REGION Network 10: Stacker General Alarm
   RUNG wire#powerrail
      { S7_Templates := "SrcType := Word" } EQ_Contact(in1 := "DB3_FAULTS".Alarm_Safety_S, in2 := 0)
      { S7_Templates := "SrcType := Word" } EQ_Contact(in1 := "DB3_FAULTS".Alarm_Safety_SN, in2 := 0)
      { S7_Templates := "SrcType := Word" } EQ_Contact(in1 := "DB3_FAULTS".Alarm_Safety_Z2, in2 := 0)
      { S7_Templates := "SrcType := Word" } EQ_Contact(in1 := "DB3_FAULTS".Alarm_Stacker, in2 := 0)
      { S7_Templates := "SrcType := Word" } EQ_Contact(in1 := "DB3_FAULTS".Alarm_General_S, in2 := 0)
      { S7_Templates := "SrcType := Word" } EQ_Contact(in1 := "DB3_FAULTS".Alarm_CD2, in2 := 0)
      { S7_Templates := "SrcType := Word" } EQ_Contact(in1 := "DB3_FAULTS".Alarm_CD1, in2 := 0)
      Coil( #NoAlmAny )
   END_RUNG
   RUNG wire#powerrail
      Contact( #NoAlmAny )
      { S7_Templates := "SrcType := Word" } EQ_Contact(in1 := "s".f[1].almw, in2 := 0)
      { S7_Templates := "SrcType := Word" } EQ_Contact(in1 := "s".f[2].almw, in2 := 0)
      { S7_Templates := "SrcType := Word" } EQ_Contact(in1 := "s".f[3].almw, in2 := 0)
      { S7_Templates := "SrcType := Word" } EQ_Contact(in1 := "s".f[4].almw, in2 := 0)
      { S7_Templates := "SrcType := Word" } EQ_Contact(in1 := "s".f[5].almw, in2 := 0)
      Coil( #NoAlmAny )
   END_RUNG
   RUNG wire#powerrail
      Contact( #NoAlmAny )
      { S7_Templates := "SrcType := Word" } EQ_Contact(in1 := "O".S_Alm_Stack_Dwn, in2 := 0)
      { S7_Templates := "SrcType := Word" } EQ_Contact(in1 := "O".S_Alm_Stack_Mid, in2 := 0)
      { S7_Templates := "SrcType := Word" } EQ_Contact(in1 := "O".S_Alm_Stack_Up, in2 := 0)
      { S7_Templates := "SrcType := Word" } EQ_Contact(in1 := "O".Centror_A.AlarmW, in2 := 0)
      { S7_Templates := "SrcType := Word" } EQ_Contact(in1 := "O".FurcaStacker.AlarmW, in2 := 0)
      I_Contact( "DB2_WORK_BITS".Stacker_Handler.Output.oAlarmForks )
      I_Contact( "DB2_WORK_BITS".Stacker_Handler.Output.oAlarmPosition )
      Coil( #NoAlmAny )
   END_RUNG
   RUNG wire#powerrail
      I_Contact( #NoAlmAny )
      I_Contact( "x"."b"[16] )
      Coil( "Gen".S_AlarmAny )
   END_RUNG
   // the same network as SCL:
   #NoAlmAny := ("DB3_FAULTS".Alarm_Safety_S = 0) AND ("DB3_FAULTS".Alarm_Safety_SN = 0) AND ("DB3_FAULTS".Alarm_Safety_Z2 = 0) AND ("DB3_FAULTS".Alarm_Stacker = 0) AND ("DB3_FAULTS".Alarm_General_S = 0) AND ("DB3_FAULTS".Alarm_CD2 = 0) AND ("DB3_FAULTS".Alarm_CD1 = 0);
   #NoAlmAny := #NoAlmAny AND ("s".f[1].almw = 0) AND ("s".f[2].almw = 0) AND ("s".f[3].almw = 0) AND ("s".f[4].almw = 0) AND ("s".f[5].almw = 0);
   #NoAlmAny := #NoAlmAny AND ("O".S_Alm_Stack_Dwn = 0) AND ("O".S_Alm_Stack_Mid = 0) AND ("O".S_Alm_Stack_Up = 0) AND ("O".Centror_A.AlarmW = 0) AND ("O".FurcaStacker.AlarmW = 0) AND NOT "DB2_WORK_BITS".Stacker_Handler.Output.oAlarmForks AND NOT "DB2_WORK_BITS".Stacker_Handler.Output.oAlarmPosition;
   "Gen".S_AlarmAny := NOT #NoAlmAny AND NOT "x"."b"[16];
END_REGION

REGION Network 11: Stacker_New General Alarm
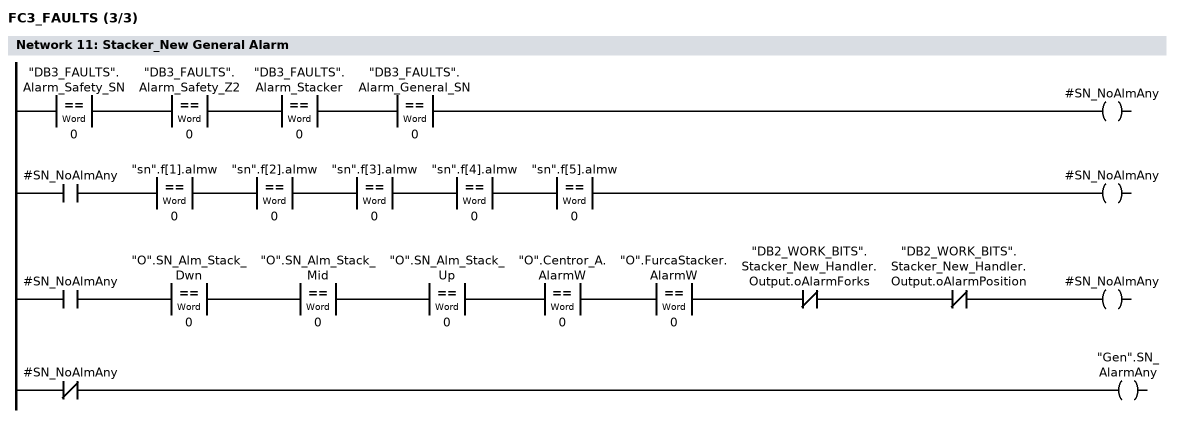
   RUNG wire#powerrail
      { S7_Templates := "SrcType := Word" } EQ_Contact(in1 := "DB3_FAULTS".Alarm_Safety_SN, in2 := 0)
      { S7_Templates := "SrcType := Word" } EQ_Contact(in1 := "DB3_FAULTS".Alarm_Safety_Z2, in2 := 0)
      { S7_Templates := "SrcType := Word" } EQ_Contact(in1 := "DB3_FAULTS".Alarm_Stacker, in2 := 0)
      { S7_Templates := "SrcType := Word" } EQ_Contact(in1 := "DB3_FAULTS".Alarm_General_SN, in2 := 0)
      Coil( #SN_NoAlmAny )
   END_RUNG
   RUNG wire#powerrail
      Contact( #SN_NoAlmAny )
      { S7_Templates := "SrcType := Word" } EQ_Contact(in1 := "sn".f[1].almw, in2 := 0)
      { S7_Templates := "SrcType := Word" } EQ_Contact(in1 := "sn".f[2].almw, in2 := 0)
      { S7_Templates := "SrcType := Word" } EQ_Contact(in1 := "sn".f[3].almw, in2 := 0)
      { S7_Templates := "SrcType := Word" } EQ_Contact(in1 := "sn".f[4].almw, in2 := 0)
      { S7_Templates := "SrcType := Word" } EQ_Contact(in1 := "sn".f[5].almw, in2 := 0)
      Coil( #SN_NoAlmAny )
   END_RUNG
   RUNG wire#powerrail
      Contact( #SN_NoAlmAny )
      { S7_Templates := "SrcType := Word" } EQ_Contact(in1 := "O".SN_Alm_Stack_Dwn, in2 := 0)
      { S7_Templates := "SrcType := Word" } EQ_Contact(in1 := "O".SN_Alm_Stack_Mid, in2 := 0)
      { S7_Templates := "SrcType := Word" } EQ_Contact(in1 := "O".SN_Alm_Stack_Up, in2 := 0)
      { S7_Templates := "SrcType := Word" } EQ_Contact(in1 := "O".Centror_A.AlarmW, in2 := 0)
      { S7_Templates := "SrcType := Word" } EQ_Contact(in1 := "O".FurcaStacker.AlarmW, in2 := 0)
      I_Contact( "DB2_WORK_BITS".Stacker_New_Handler.Output.oAlarmForks )
      I_Contact( "DB2_WORK_BITS".Stacker_New_Handler.Output.oAlarmPosition )
      Coil( #SN_NoAlmAny )
   END_RUNG
   RUNG wire#powerrail
      I_Contact( #SN_NoAlmAny )
      Coil( "Gen".SN_AlarmAny )
   END_RUNG
   // the same network as SCL:
   #SN_NoAlmAny := ("DB3_FAULTS".Alarm_Safety_SN = 0) AND ("DB3_FAULTS".Alarm_Safety_Z2 = 0) AND ("DB3_FAULTS".Alarm_Stacker = 0) AND ("DB3_FAULTS".Alarm_General_SN = 0);
   #SN_NoAlmAny := #SN_NoAlmAny AND ("sn".f[1].almw = 0) AND ("sn".f[2].almw = 0) AND ("sn".f[3].almw = 0) AND ("sn".f[4].almw = 0) AND ("sn".f[5].almw = 0);
   #SN_NoAlmAny := #SN_NoAlmAny AND ("O".SN_Alm_Stack_Dwn = 0) AND ("O".SN_Alm_Stack_Mid = 0) AND ("O".SN_Alm_Stack_Up = 0) AND ("O".Centror_A.AlarmW = 0) AND ("O".FurcaStacker.AlarmW = 0) AND NOT "DB2_WORK_BITS".Stacker_New_Handler.Output.oAlarmForks AND NOT "DB2_WORK_BITS".Stacker_New_Handler.Output.oAlarmPosition;
   "Gen".SN_AlarmAny := NOT #SN_NoAlmAny;
END_REGION
END_FUNCTION

FUNCTION "FC6_OUTPUTS" : Void   // FC6, LAD
{ S7_Optimized_Access := 'TRUE' }
VERSION : 0.1
   VAR_TEMP
      S_bsy : Bool;
      S_bsg : Bool;
      S_bsr : Bool;
      S_bsgc : Bool;
      cfo1 : Bool;
      cfo2 : Bool;
      cfo3 : Bool;
      cfA : Bool;
      SN_bsr : Bool;
      SN_bsy : Bool;
      SN_bsgc : Bool;
      SN_bsg : Bool;
      SN_cfo1 : Bool;
      SN_cfo2 : Bool;
      SN_cfo3 : Bool;
      SN_cfA : Bool;
   END_VAR
   VAR_TEMP   // added for the SCL form of the ladder/FBD networks
      _w1 : Bool;
   END_VAR
BEGIN

REGION Network 1: Stacking_New VFD Input Conveyor
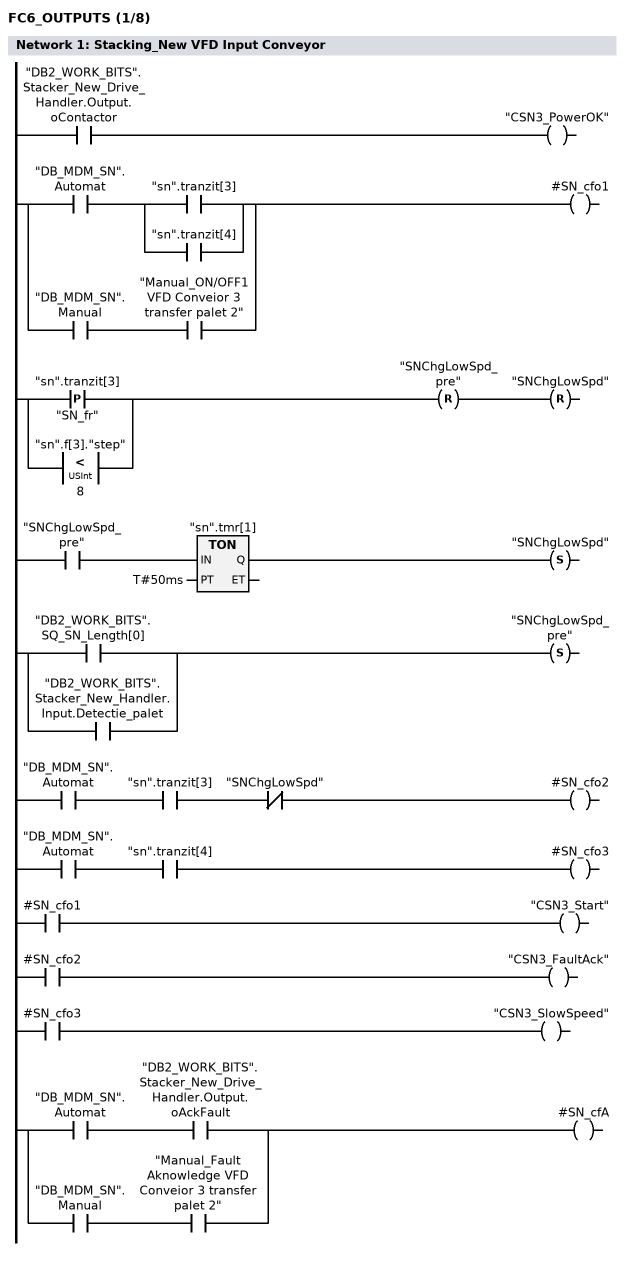
   "CSN3_PowerOK" := "DB2_WORK_BITS".Stacker_New_Drive_Handler.Output.oContactor;
   #SN_cfo1 := ("DB_MDM_SN".Automat AND ("sn".tranzit[3] OR "sn".tranzit[4])) OR ("DB_MDM_SN".Manual AND "Manual_ON/OFF1 VFD Conveior 3 transfer palet 2");
   #_w1 := "sn".tranzit[3] AND NOT "SN_fr";   // rising edge of "sn".tranzit[3]
   "SN_fr" := "sn".tranzit[3];
   IF #_w1 OR ("sn".f[3]."step" < 8) THEN
       "SNChgLowSpd_pre" := FALSE;
       "SNChgLowSpd" := FALSE;
   END_IF;
   "sn".tmr[1].TON(IN := "SNChgLowSpd_pre", PT := T#50ms);
   IF "sn".tmr[1].Q THEN "SNChgLowSpd" := TRUE; END_IF;
   IF "DB2_WORK_BITS".SQ_SN_Length[0] OR "DB2_WORK_BITS".Stacker_New_Handler.Input.Detectie_palet THEN
       "SNChgLowSpd_pre" := TRUE;
   END_IF;
   #SN_cfo2 := "DB_MDM_SN".Automat AND "sn".tranzit[3] AND NOT "SNChgLowSpd";
   #SN_cfo3 := "DB_MDM_SN".Automat AND "sn".tranzit[4];
   "CSN3_Start" := #SN_cfo1;
   "CSN3_FaultAck" := #SN_cfo2;
   "CSN3_SlowSpeed" := #SN_cfo3;
   #SN_cfA := ("DB_MDM_SN".Automat AND "DB2_WORK_BITS".Stacker_New_Drive_Handler.Output.oAckFault) OR ("DB_MDM_SN".Manual AND "Manual_Fault Aknowledge VFD Conveior 3 transfer palet 2");
END_REGION

REGION Network 2: Stacking_New VFD Output Conveyor
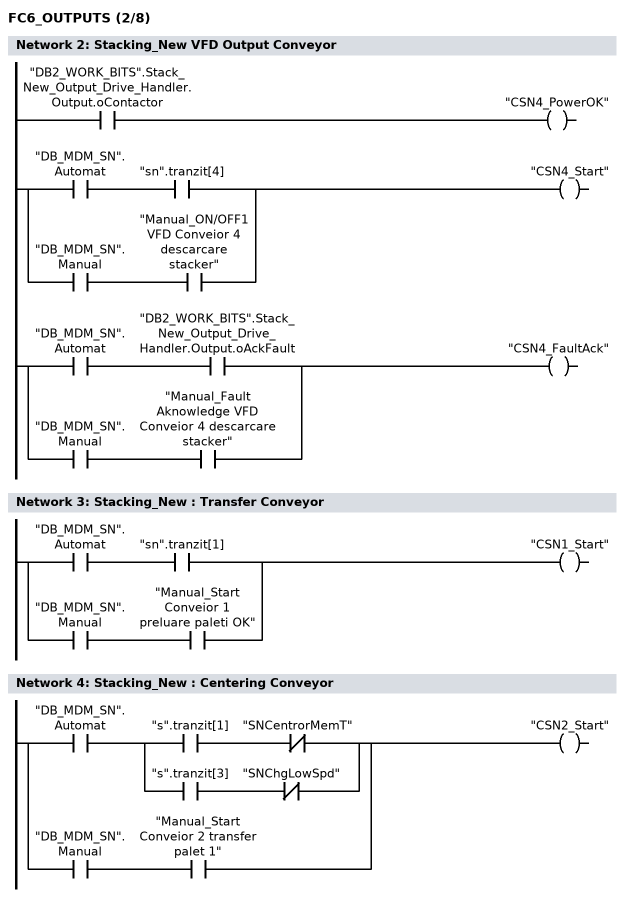
   RUNG wire#powerrail
      Contact( "DB2_WORK_BITS".Stack_New_Output_Drive_Handler.Output.oContactor )
      Coil( "CSN4_PowerOK" )
   END_RUNG
   RUNG wire#powerrail
      Contact( "DB_MDM_SN".Automat )
      Contact( "sn".tranzit[4] )
      wire#w1
      Coil( "CSN4_Start" )
   END_RUNG
   RUNG wire#powerrail
      Contact( "DB_MDM_SN".Manual )
      Contact( "Manual_ON/OFF1 VFD Conveior 4 descarcare stacker" )
   END_RUNG wire#w1
   RUNG wire#powerrail
      Contact( "DB_MDM_SN".Automat )
      Contact( "DB2_WORK_BITS".Stack_New_Output_Drive_Handler.Output.oAckFault )
      wire#w2
      Coil( "CSN4_FaultAck" )
   END_RUNG
   RUNG wire#powerrail
      Contact( "DB_MDM_SN".Manual )
      Contact( "Manual_Fault Aknowledge VFD Conveior 4 descarcare stacker" )
   END_RUNG wire#w2
   // the same network as SCL:
   "CSN4_PowerOK" := "DB2_WORK_BITS".Stack_New_Output_Drive_Handler.Output.oContactor;
   "CSN4_Start" := ("DB_MDM_SN".Automat AND "sn".tranzit[4]) OR ("DB_MDM_SN".Manual AND "Manual_ON/OFF1 VFD Conveior 4 descarcare stacker");
   "CSN4_FaultAck" := ("DB_MDM_SN".Automat AND "DB2_WORK_BITS".Stack_New_Output_Drive_Handler.Output.oAckFault) OR ("DB_MDM_SN".Manual AND "Manual_Fault Aknowledge VFD Conveior 4 descarcare stacker");
END_REGION

REGION Network 3: Stacking_New : Transfer Conveyor
   RUNG wire#powerrail
      Contact( "DB_MDM_SN".Automat )
      Contact( "sn".tranzit[1] )
      wire#w1
      Coil( "CSN1_Start" )
   END_RUNG
   RUNG wire#powerrail
      Contact( "DB_MDM_SN".Manual )
      Contact( "Manual_Start Conveior 1 preluare paleti OK" )
   END_RUNG wire#w1
   // the same network as SCL:
   "CSN1_Start" := ("DB_MDM_SN".Automat AND "sn".tranzit[1]) OR ("DB_MDM_SN".Manual AND "Manual_Start Conveior 1 preluare paleti OK");
END_REGION

REGION Network 4: Stacking_New : Centering Conveyor
   RUNG wire#powerrail
      Contact( "DB_MDM_SN".Automat )
      wire#w1
      Contact( "s".tranzit[1] )
      I_Contact( "SNCentrorMemT" )
      wire#w2
      Coil( "CSN2_Start" )
   END_RUNG
   RUNG wire#w1
      Contact( "s".tranzit[3] )
      I_Contact( "SNChgLowSpd" )
   END_RUNG wire#w2
   RUNG wire#powerrail
      Contact( "DB_MDM_SN".Manual )
      Contact( "Manual_Start Conveior 2 transfer palet 1" )
   END_RUNG wire#w2
   // the same network as SCL:
   "CSN2_Start" := ("DB_MDM_SN".Automat AND (("s".tranzit[1] AND NOT "SNCentrorMemT") OR ("s".tranzit[3] AND NOT "SNChgLowSpd"))) OR ("DB_MDM_SN".Manual AND "Manual_Start Conveior 2 transfer palet 1");
END_REGION

REGION Network 5: Stacking : VFD Input Conveyor
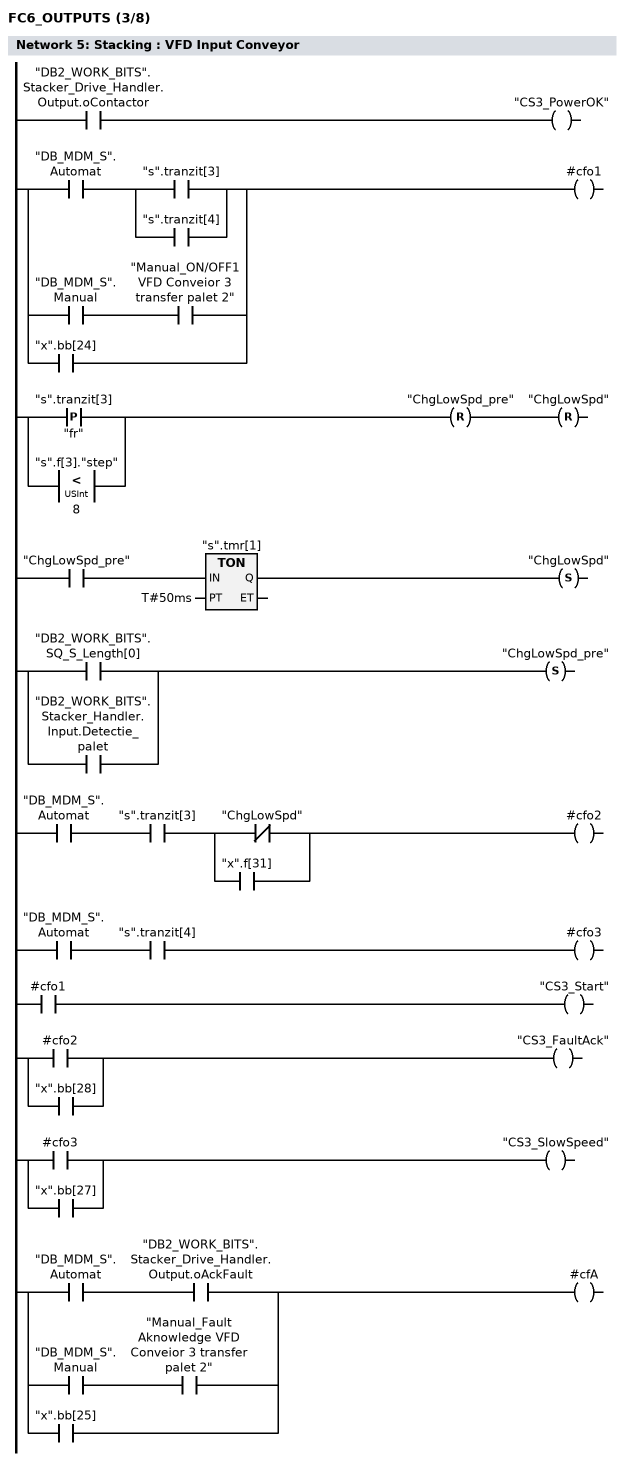
   "CS3_PowerOK" := "DB2_WORK_BITS".Stacker_Drive_Handler.Output.oContactor;
   #cfo1 := ("DB_MDM_S".Automat AND ("s".tranzit[3] OR "s".tranzit[4])) OR ("DB_MDM_S".Manual AND "Manual_ON/OFF1 VFD Conveior 3 transfer palet 2") OR "x".bb[24];
   #_w1 := "s".tranzit[3] AND NOT "fr";   // rising edge of "s".tranzit[3]
   "fr" := "s".tranzit[3];
   IF #_w1 OR ("s".f[3]."step" < 8) THEN
       "ChgLowSpd_pre" := FALSE;
       "ChgLowSpd" := FALSE;
   END_IF;
   "s".tmr[1].TON(IN := "ChgLowSpd_pre", PT := T#50ms);
   IF "s".tmr[1].Q THEN "ChgLowSpd" := TRUE; END_IF;
   IF "DB2_WORK_BITS".SQ_S_Length[0] OR "DB2_WORK_BITS".Stacker_Handler.Input.Detectie_palet THEN
       "ChgLowSpd_pre" := TRUE;
   END_IF;
   #cfo2 := "DB_MDM_S".Automat AND "s".tranzit[3] AND (NOT "ChgLowSpd" OR "x".f[31]);
   #cfo3 := "DB_MDM_S".Automat AND "s".tranzit[4];
   "CS3_Start" := #cfo1;
   "CS3_FaultAck" := #cfo2 OR "x".bb[28];
   "CS3_SlowSpeed" := #cfo3 OR "x".bb[27];
   #cfA := ("DB_MDM_S".Automat AND "DB2_WORK_BITS".Stacker_Drive_Handler.Output.oAckFault) OR ("DB_MDM_S".Manual AND "Manual_Fault Aknowledge VFD Conveior 3 transfer palet 2") OR "x".bb[25];
END_REGION

REGION Network 6: Stacking : VFD Output Conveyor
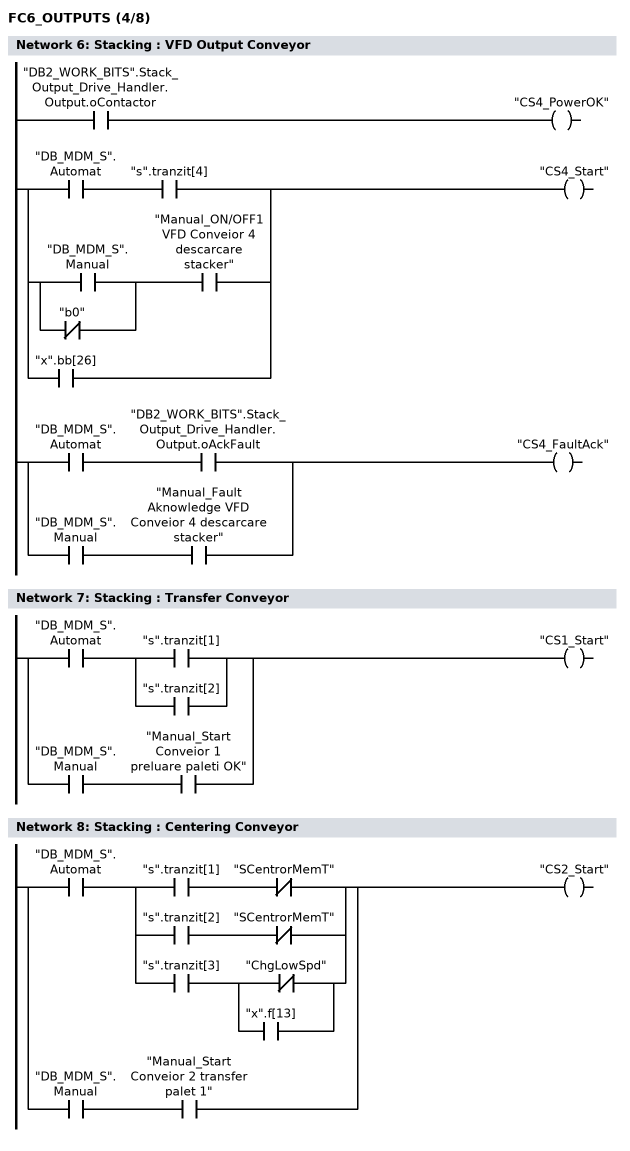
   RUNG wire#powerrail
      Contact( "DB2_WORK_BITS".Stack_Output_Drive_Handler.Output.oContactor )
      Coil( "CS4_PowerOK" )
   END_RUNG
   RUNG wire#powerrail
      Contact( "DB_MDM_S".Automat )
      Contact( "s".tranzit[4] )
      wire#w1
      Coil( "CS4_Start" )
   END_RUNG
   RUNG wire#powerrail
      Contact( "DB_MDM_S".Manual )
      wire#w2
      Contact( "Manual_ON/OFF1 VFD Conveior 4 descarcare stacker" )
   END_RUNG wire#w1
   RUNG wire#powerrail
      I_Contact( "b0" )
   END_RUNG wire#w2
   RUNG wire#powerrail
      Contact( "x".bb[26] )
   END_RUNG wire#w1
   RUNG wire#powerrail
      Contact( "DB_MDM_S".Automat )
      Contact( "DB2_WORK_BITS".Stack_Output_Drive_Handler.Output.oAckFault )
      wire#w3
      Coil( "CS4_FaultAck" )
   END_RUNG
   RUNG wire#powerrail
      Contact( "DB_MDM_S".Manual )
      Contact( "Manual_Fault Aknowledge VFD Conveior 4 descarcare stacker" )
   END_RUNG wire#w3
   // the same network as SCL:
   "CS4_PowerOK" := "DB2_WORK_BITS".Stack_Output_Drive_Handler.Output.oContactor;
   "CS4_Start" := ("DB_MDM_S".Automat AND "s".tranzit[4]) OR (("DB_MDM_S".Manual OR NOT "b0") AND "Manual_ON/OFF1 VFD Conveior 4 descarcare stacker") OR "x".bb[26];
   "CS4_FaultAck" := ("DB_MDM_S".Automat AND "DB2_WORK_BITS".Stack_Output_Drive_Handler.Output.oAckFault) OR ("DB_MDM_S".Manual AND "Manual_Fault Aknowledge VFD Conveior 4 descarcare stacker");
END_REGION

REGION Network 7: Stacking : Transfer Conveyor
   RUNG wire#powerrail
      Contact( "DB_MDM_S".Automat )
      wire#w1
      Contact( "s".tranzit[1] )
      wire#w2
      Coil( "CS1_Start" )
   END_RUNG
   RUNG wire#w1
      Contact( "s".tranzit[2] )
   END_RUNG wire#w2
   RUNG wire#powerrail
      Contact( "DB_MDM_S".Manual )
      Contact( "Manual_Start Conveior 1 preluare paleti OK" )
   END_RUNG wire#w2
   // the same network as SCL:
   "CS1_Start" := ("DB_MDM_S".Automat AND ("s".tranzit[1] OR "s".tranzit[2])) OR ("DB_MDM_S".Manual AND "Manual_Start Conveior 1 preluare paleti OK");
END_REGION

REGION Network 8: Stacking : Centering Conveyor
   RUNG wire#powerrail
      Contact( "DB_MDM_S".Automat )
      wire#w1
      Contact( "s".tranzit[1] )
      I_Contact( "SCentrorMemT" )
      wire#w2
      Coil( "CS2_Start" )
   END_RUNG
   RUNG wire#w1
      Contact( "s".tranzit[2] )
      I_Contact( "SCentrorMemT" )
   END_RUNG wire#w2
   RUNG wire#w1
      Contact( "s".tranzit[3] )
      wire#w3
      I_Contact( "ChgLowSpd" )
   END_RUNG wire#w2
   RUNG wire#w3
      Contact( "x".f[13] )
   END_RUNG wire#w2
   RUNG wire#powerrail
      Contact( "DB_MDM_S".Manual )
      Contact( "Manual_Start Conveior 2 transfer palet 1" )
   END_RUNG wire#w2
   // the same network as SCL:
   "CS2_Start" := ("DB_MDM_S".Automat AND (("s".tranzit[1] AND NOT "SCentrorMemT") OR ("s".tranzit[2] AND NOT "SCentrorMemT") OR ("s".tranzit[3] AND (NOT "ChgLowSpd" OR "x".f[13])))) OR ("DB_MDM_S".Manual AND "Manual_Start Conveior 2 transfer palet 1");
END_REGION

REGION Network 9: Stacking_New : Comanda SoftStart Power ON
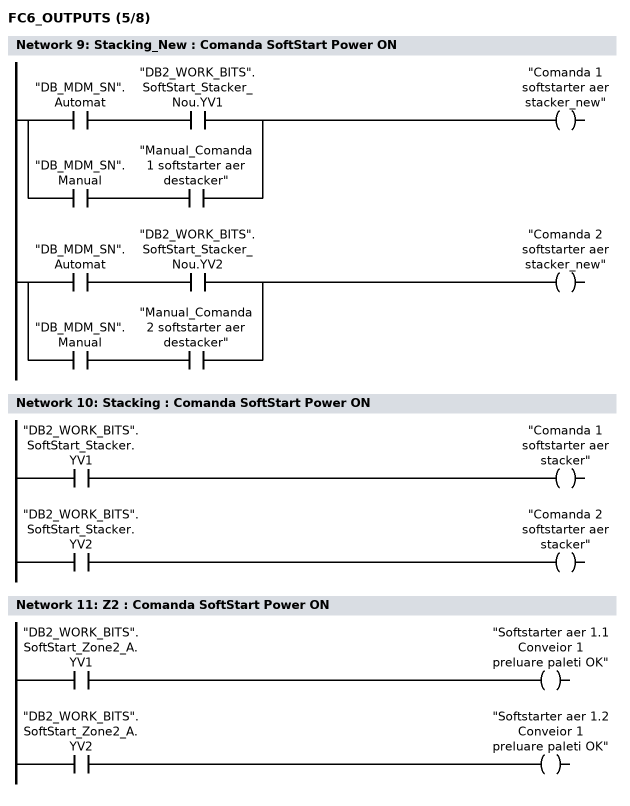
   RUNG wire#powerrail
      Contact( "DB_MDM_SN".Automat )
      Contact( "DB2_WORK_BITS".SoftStart_Stacker_Nou.YV1 )
      wire#w1
      Coil( "Comanda 1 softstarter aer stacker_new" )
   END_RUNG
   RUNG wire#powerrail
      Contact( "DB_MDM_SN".Manual )
      Contact( "Manual_Comanda 1 softstarter aer destacker" )
   END_RUNG wire#w1
   RUNG wire#powerrail
      Contact( "DB_MDM_SN".Automat )
      Contact( "DB2_WORK_BITS".SoftStart_Stacker_Nou.YV2 )
      wire#w2
      Coil( "Comanda 2 softstarter aer stacker_new" )
   END_RUNG
   RUNG wire#powerrail
      Contact( "DB_MDM_SN".Manual )
      Contact( "Manual_Comanda 2 softstarter aer destacker" )
   END_RUNG wire#w2
   // the same network as SCL:
   "Comanda 1 softstarter aer stacker_new" := ("DB_MDM_SN".Automat AND "DB2_WORK_BITS".SoftStart_Stacker_Nou.YV1) OR ("DB_MDM_SN".Manual AND "Manual_Comanda 1 softstarter aer destacker");
   "Comanda 2 softstarter aer stacker_new" := ("DB_MDM_SN".Automat AND "DB2_WORK_BITS".SoftStart_Stacker_Nou.YV2) OR ("DB_MDM_SN".Manual AND "Manual_Comanda 2 softstarter aer destacker");
END_REGION

REGION Network 10: Stacking : Comanda SoftStart Power ON
   RUNG wire#powerrail
      Contact( "DB2_WORK_BITS".SoftStart_Stacker.YV1 )
      Coil( "Comanda 1 softstarter aer stacker" )
   END_RUNG
   RUNG wire#powerrail
      Contact( "DB2_WORK_BITS".SoftStart_Stacker.YV2 )
      Coil( "Comanda 2 softstarter aer stacker" )
   END_RUNG
   // the same network as SCL:
   "Comanda 1 softstarter aer stacker" := "DB2_WORK_BITS".SoftStart_Stacker.YV1;
   "Comanda 2 softstarter aer stacker" := "DB2_WORK_BITS".SoftStart_Stacker.YV2;
END_REGION

REGION Network 11: Z2 : Comanda SoftStart Power ON
   RUNG wire#powerrail
      Contact( "DB2_WORK_BITS".SoftStart_Zone2_A.YV1 )
      Coil( "Softstarter aer 1.1 Conveior 1 preluare paleti OK" )
   END_RUNG
   RUNG wire#powerrail
      Contact( "DB2_WORK_BITS".SoftStart_Zone2_A.YV2 )
      Coil( "Softstarter aer 1.2 Conveior 1 preluare paleti OK" )
   END_RUNG
   // the same network as SCL:
   "Softstarter aer 1.1 Conveior 1 preluare paleti OK" := "DB2_WORK_BITS".SoftStart_Zone2_A.YV1;
   "Softstarter aer 1.2 Conveior 1 preluare paleti OK" := "DB2_WORK_BITS".SoftStart_Zone2_A.YV2;
END_REGION

REGION Network 12: Rearm safety
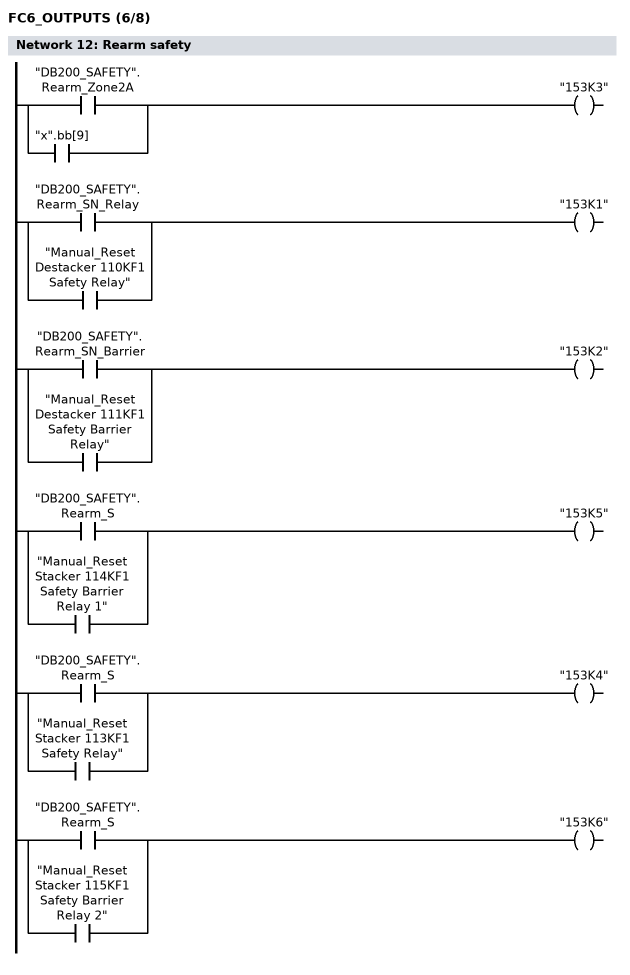
   RUNG wire#powerrail
      Contact( "DB200_SAFETY".Rearm_Zone2A )
      wire#w1
      Coil( "153K3" )
   END_RUNG
   RUNG wire#powerrail
      Contact( "x".bb[9] )
   END_RUNG wire#w1
   RUNG wire#powerrail
      Contact( "DB200_SAFETY".Rearm_SN_Relay )
      wire#w2
      Coil( "153K1" )
   END_RUNG
   RUNG wire#powerrail
      Contact( "Manual_Reset Destacker 110KF1 Safety Relay" )
   END_RUNG wire#w2
   RUNG wire#powerrail
      Contact( "DB200_SAFETY".Rearm_SN_Barrier )
      wire#w3
      Coil( "153K2" )
   END_RUNG
   RUNG wire#powerrail
      Contact( "Manual_Reset Destacker 111KF1 Safety Barrier Relay" )
   END_RUNG wire#w3
   RUNG wire#powerrail
      Contact( "DB200_SAFETY".Rearm_S )
      wire#w4
      Coil( "153K5" )
   END_RUNG
   RUNG wire#powerrail
      Contact( "Manual_Reset Stacker 114KF1 Safety Barrier Relay 1" )
   END_RUNG wire#w4
   RUNG wire#powerrail
      Contact( "DB200_SAFETY".Rearm_S )
      wire#w5
      Coil( "153K4" )
   END_RUNG
   RUNG wire#powerrail
      Contact( "Manual_Reset Stacker 113KF1 Safety Relay" )
   END_RUNG wire#w5
   RUNG wire#powerrail
      Contact( "DB200_SAFETY".Rearm_S )
      wire#w6
      Coil( "153K6" )
   END_RUNG
   RUNG wire#powerrail
      Contact( "Manual_Reset Stacker 115KF1 Safety Barrier Relay 2" )
   END_RUNG wire#w6
   // the same network as SCL:
   "153K3" := "DB200_SAFETY".Rearm_Zone2A OR "x".bb[9];
   "153K1" := "DB200_SAFETY".Rearm_SN_Relay OR "Manual_Reset Destacker 110KF1 Safety Relay";
   "153K2" := "DB200_SAFETY".Rearm_SN_Barrier OR "Manual_Reset Destacker 111KF1 Safety Barrier Relay";
   "153K5" := "DB200_SAFETY".Rearm_S OR "Manual_Reset Stacker 114KF1 Safety Barrier Relay 1";
   "153K4" := "DB200_SAFETY".Rearm_S OR "Manual_Reset Stacker 113KF1 Safety Relay";
   "153K6" := "DB200_SAFETY".Rearm_S OR "Manual_Reset Stacker 115KF1 Safety Barrier Relay 2";
END_REGION

REGION Network 13: Stacking : Control Balize
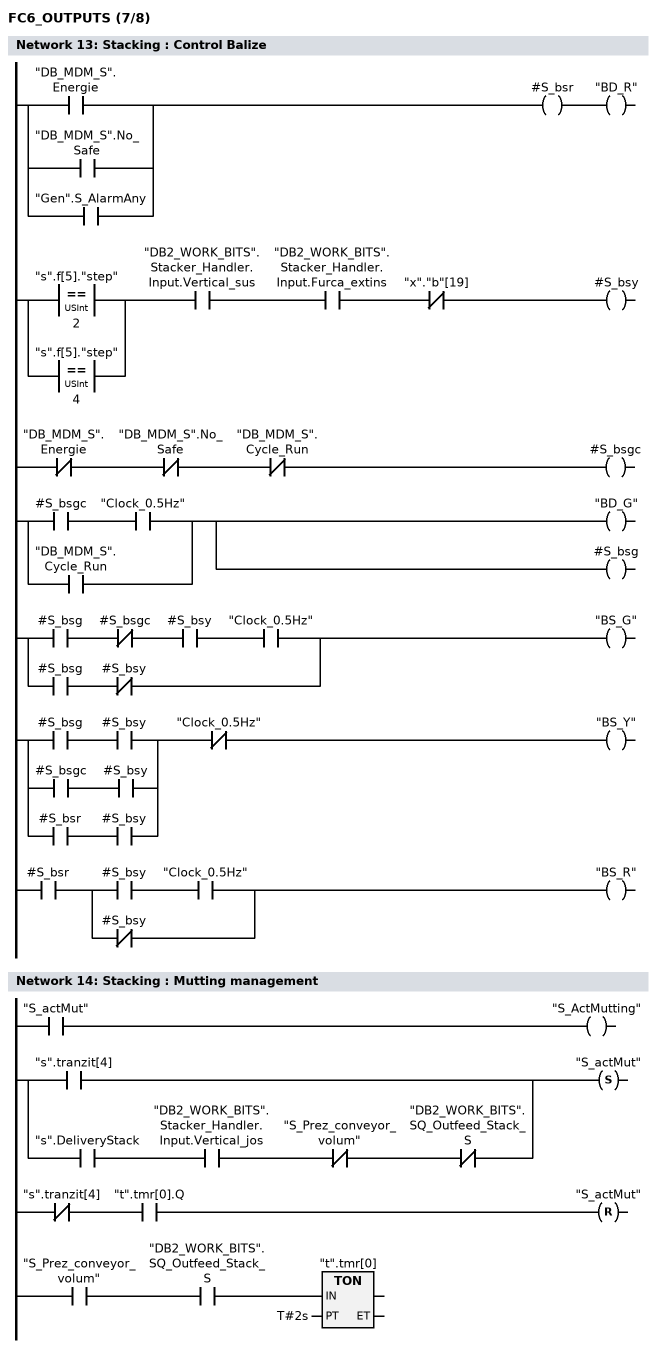
   RUNG wire#powerrail
      Contact( "DB_MDM_S".Energie )
      wire#w1
      Coil( #S_bsr )
      Coil( "BD_R" )
   END_RUNG
   RUNG wire#powerrail
      Contact( "DB_MDM_S".No_Safe )
   END_RUNG wire#w1
   RUNG wire#powerrail
      Contact( "Gen".S_AlarmAny )
   END_RUNG wire#w1
   RUNG wire#powerrail
      { S7_Templates := "SrcType := USInt" } EQ_Contact(in1 := "s".f[5]."step", in2 := 2)
      wire#w2
      Contact( "DB2_WORK_BITS".Stacker_Handler.Input.Vertical_sus )
      Contact( "DB2_WORK_BITS".Stacker_Handler.Input.Furca_extins )
      I_Contact( "x"."b"[19] )
      Coil( #S_bsy )
   END_RUNG
   RUNG wire#powerrail
      { S7_Templates := "SrcType := USInt" } EQ_Contact(in1 := "s".f[5]."step", in2 := 4)
   END_RUNG wire#w2
   RUNG wire#powerrail
      I_Contact( "DB_MDM_S".Energie )
      I_Contact( "DB_MDM_S".No_Safe )
      I_Contact( "DB_MDM_S".Cycle_Run )
      Coil( #S_bsgc )
   END_RUNG
   RUNG wire#powerrail
      Contact( #S_bsgc )
      Contact( "Clock_0.5Hz" )
      wire#w3
      Coil( "BD_G" )
   END_RUNG
   RUNG wire#powerrail
      Contact( "DB_MDM_S".Cycle_Run )
   END_RUNG wire#w3
   RUNG wire#w3
      Coil( #S_bsg )
   END_RUNG
   RUNG wire#powerrail
      Contact( #S_bsg )
      I_Contact( #S_bsgc )
      Contact( #S_bsy )
      Contact( "Clock_0.5Hz" )
      wire#w4
      Coil( "BS_G" )
   END_RUNG
   RUNG wire#powerrail
      Contact( #S_bsg )
      I_Contact( #S_bsy )
   END_RUNG wire#w4
   RUNG wire#powerrail
      Contact( #S_bsg )
      Contact( #S_bsy )
      wire#w5
      I_Contact( "Clock_0.5Hz" )
      Coil( "BS_Y" )
   END_RUNG
   RUNG wire#powerrail
      Contact( #S_bsgc )
      Contact( #S_bsy )
   END_RUNG wire#w5
   RUNG wire#powerrail
      Contact( #S_bsr )
      Contact( #S_bsy )
   END_RUNG wire#w5
   RUNG wire#powerrail
      Contact( #S_bsr )
      wire#w6
      Contact( #S_bsy )
      Contact( "Clock_0.5Hz" )
      wire#w7
      Coil( "BS_R" )
   END_RUNG
   RUNG wire#w6
      I_Contact( #S_bsy )
   END_RUNG wire#w7
   // the same network as SCL:
   #S_bsr := "DB_MDM_S".Energie OR "DB_MDM_S".No_Safe OR "Gen".S_AlarmAny;
   "BD_R" := #S_bsr;
   #S_bsy := (("s".f[5]."step" = 2) OR ("s".f[5]."step" = 4)) AND "DB2_WORK_BITS".Stacker_Handler.Input.Vertical_sus AND "DB2_WORK_BITS".Stacker_Handler.Input.Furca_extins AND NOT "x"."b"[19];
   #S_bsgc := NOT "DB_MDM_S".Energie AND NOT "DB_MDM_S".No_Safe AND NOT "DB_MDM_S".Cycle_Run;
   "BD_G" := (#S_bsgc AND "Clock_0.5Hz") OR "DB_MDM_S".Cycle_Run;
   #S_bsg := "BD_G";
   "BS_G" := (#S_bsg AND NOT #S_bsgc AND #S_bsy AND "Clock_0.5Hz") OR (#S_bsg AND NOT #S_bsy);
   "BS_Y" := ((#S_bsg AND #S_bsy) OR (#S_bsgc AND #S_bsy) OR (#S_bsr AND #S_bsy)) AND NOT "Clock_0.5Hz";
   "BS_R" := #S_bsr AND ((#S_bsy AND "Clock_0.5Hz") OR NOT #S_bsy);
END_REGION

REGION Network 14: Stacking : Mutting management
   "S_ActMutting" := "S_actMut";
   IF "s".tranzit[4] OR ("s".DeliveryStack AND "DB2_WORK_BITS".Stacker_Handler.Input.Vertical_jos AND NOT "S_Prez_conveyor_volum" AND NOT "DB2_WORK_BITS".SQ_Outfeed_Stack_S) THEN
       "S_actMut" := TRUE;
   END_IF;
   IF NOT "s".tranzit[4] AND "t".tmr[0].Q THEN "S_actMut" := FALSE; END_IF;
   "t".tmr[0].TON(IN := "S_Prez_conveyor_volum" AND "DB2_WORK_BITS".SQ_Outfeed_Stack_S, PT := T#2s);
END_REGION

REGION Network 15: Stacking_New : Mutting management
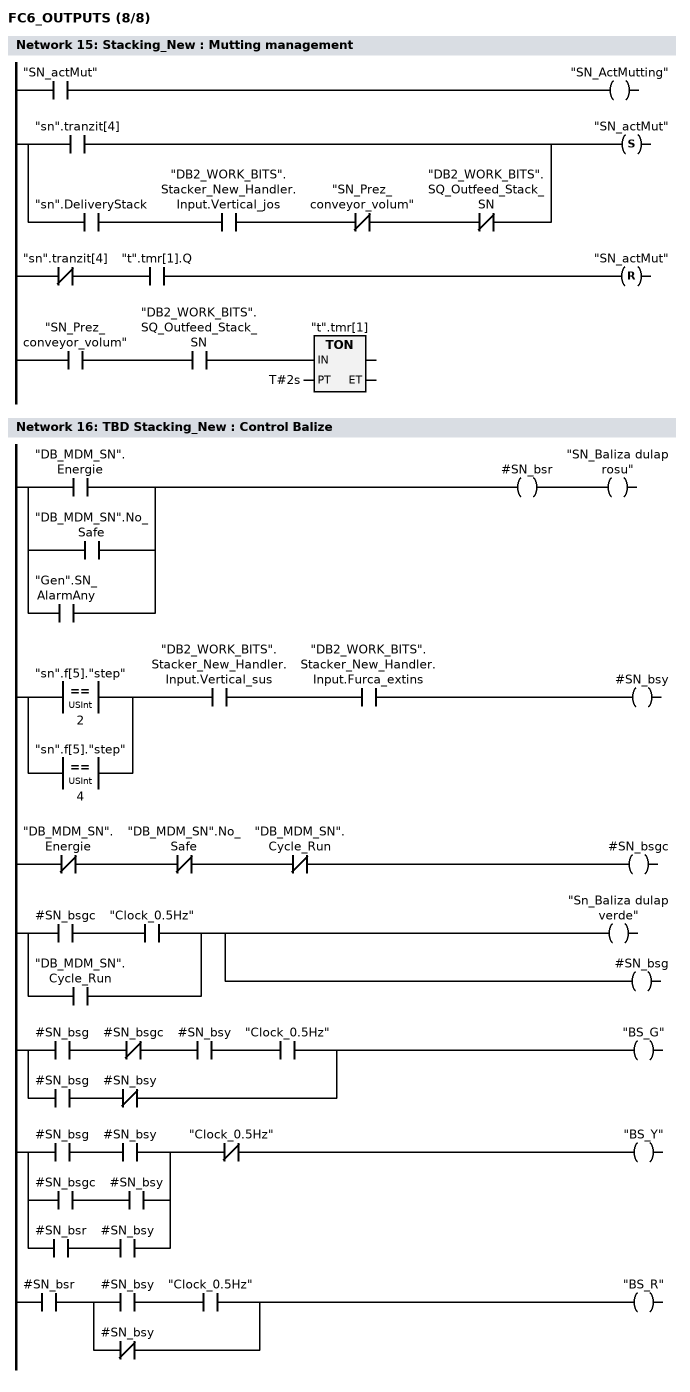
   "SN_ActMutting" := "SN_actMut";
   IF "sn".tranzit[4] OR ("sn".DeliveryStack AND "DB2_WORK_BITS".Stacker_New_Handler.Input.Vertical_jos AND NOT "SN_Prez_conveyor_volum" AND NOT "DB2_WORK_BITS".SQ_Outfeed_Stack_SN) THEN
       "SN_actMut" := TRUE;
   END_IF;
   IF NOT "sn".tranzit[4] AND "t".tmr[1].Q THEN "SN_actMut" := FALSE; END_IF;
   "t".tmr[1].TON(IN := "SN_Prez_conveyor_volum" AND "DB2_WORK_BITS".SQ_Outfeed_Stack_SN, PT := T#2s);
END_REGION
